REGION Network 203: DB64 DBX44.7 = PVVA Tank 8 Open Alarm
   // BWTS_ALARM_WORD_23_BIT_7
   RUNG wire#powerrail
      Contact( "1092_HMI_OP_FLAGS".CV427_428_PVVA_Alarms[8].Open )
      Coil( %DB60.DBX44.7 )
   END_RUNG
   // the same network as SCL:
   %DB60.DBX44.7 := "1092_HMI_OP_FLAGS".CV427_428_PVVA_Alarms[8].Open;
END_REGION

REGION Network 204: DB64 DBX45.0 = PVVA Tank 9 Open Alarm
   // BWTS_ALARM_WORD_23_BIT_8
   RUNG wire#powerrail
      Contact( "1092_HMI_OP_FLAGS".CV427_428_PVVA_Alarms[9].Open )
      Coil( %DB60.DBX45.0 )
   END_RUNG
   // the same network as SCL:
   %DB60.DBX45.0 := "1092_HMI_OP_FLAGS".CV427_428_PVVA_Alarms[9].Open;
END_REGION

REGION Network 205: DB64 DBX45.1 = PVVA Tank 10 Open Alarm
   // BWTS_ALARM_WORD_23_BIT_9
   RUNG wire#powerrail
      Contact( "1092_HMI_OP_FLAGS".CV427_428_PVVA_Alarms[10].Open )
      Coil( %DB60.DBX45.1 )
   END_RUNG
   // the same network as SCL:
   %DB60.DBX45.1 := "1092_HMI_OP_FLAGS".CV427_428_PVVA_Alarms[10].Open;
END_REGION

REGION Network 206: DB64 DBX45.2 = PVVA Tank 11 Open Alarm
   // BWTS_ALARM_WORD_23_BIT_10
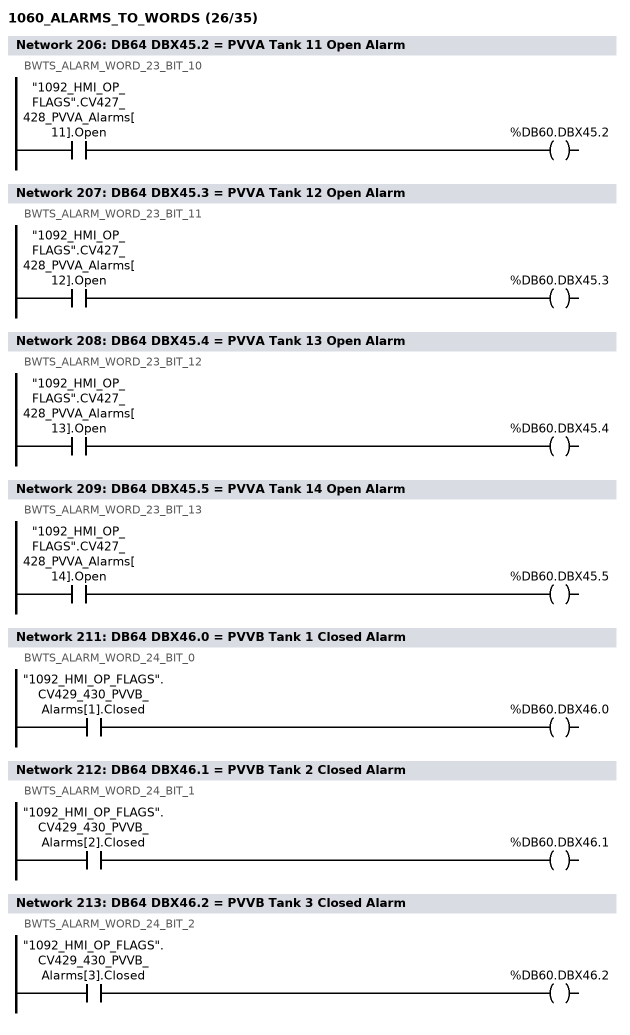
   RUNG wire#powerrail
      Contact( "1092_HMI_OP_FLAGS".CV427_428_PVVA_Alarms[11].Open )
      Coil( %DB60.DBX45.2 )
   END_RUNG
   // the same network as SCL:
   %DB60.DBX45.2 := "1092_HMI_OP_FLAGS".CV427_428_PVVA_Alarms[11].Open;
END_REGION

REGION Network 207: DB64 DBX45.3 = PVVA Tank 12 Open Alarm
   // BWTS_ALARM_WORD_23_BIT_11
   RUNG wire#powerrail
      Contact( "1092_HMI_OP_FLAGS".CV427_428_PVVA_Alarms[12].Open )
      Coil( %DB60.DBX45.3 )
   END_RUNG
   // the same network as SCL:
   %DB60.DBX45.3 := "1092_HMI_OP_FLAGS".CV427_428_PVVA_Alarms[12].Open;
END_REGION

REGION Network 208: DB64 DBX45.4 = PVVA Tank 13 Open Alarm
   // BWTS_ALARM_WORD_23_BIT_12
   RUNG wire#powerrail
      Contact( "1092_HMI_OP_FLAGS".CV427_428_PVVA_Alarms[13].Open )
      Coil( %DB60.DBX45.4 )
   END_RUNG
   // the same network as SCL:
   %DB60.DBX45.4 := "1092_HMI_OP_FLAGS".CV427_428_PVVA_Alarms[13].Open;
END_REGION

REGION Network 209: DB64 DBX45.5 = PVVA Tank 14 Open Alarm
   // BWTS_ALARM_WORD_23_BIT_13
   RUNG wire#powerrail
      Contact( "1092_HMI_OP_FLAGS".CV427_428_PVVA_Alarms[14].Open )
      Coil( %DB60.DBX45.5 )
   END_RUNG
   // the same network as SCL:
   %DB60.DBX45.5 := "1092_HMI_OP_FLAGS".CV427_428_PVVA_Alarms[14].Open;
END_REGION

REGION Network 211: DB64 DBX46.0 = PVVB Tank 1 Closed Alarm
   // BWTS_ALARM_WORD_24_BIT_0
   RUNG wire#powerrail
      Contact( "1092_HMI_OP_FLAGS".CV429_430_PVVB_Alarms[1].Closed )
      Coil( %DB60.DBX46.0 )
   END_RUNG
   // the same network as SCL:
   %DB60.DBX46.0 := "1092_HMI_OP_FLAGS".CV429_430_PVVB_Alarms[1].Closed;
END_REGION

REGION Network 212: DB64 DBX46.1 = PVVB Tank 2 Closed Alarm
   // BWTS_ALARM_WORD_24_BIT_1
   RUNG wire#powerrail
      Contact( "1092_HMI_OP_FLAGS".CV429_430_PVVB_Alarms[2].Closed )
      Coil( %DB60.DBX46.1 )
   END_RUNG
   // the same network as SCL:
   %DB60.DBX46.1 := "1092_HMI_OP_FLAGS".CV429_430_PVVB_Alarms[2].Closed;
END_REGION

REGION Network 213: DB64 DBX46.2 = PVVB Tank 3 Closed Alarm
   // BWTS_ALARM_WORD_24_BIT_2
   RUNG wire#powerrail
      Contact( "1092_HMI_OP_FLAGS".CV429_430_PVVB_Alarms[3].Closed )
      Coil( %DB60.DBX46.2 )
   END_RUNG
   // the same network as SCL:
   %DB60.DBX46.2 := "1092_HMI_OP_FLAGS".CV429_430_PVVB_Alarms[3].Closed;
END_REGION

REGION Network 214: DB64 DBX46.3 = PVVB Tank 4 Closed Alarm
   // BWTS_ALARM_WORD_24_BIT_3
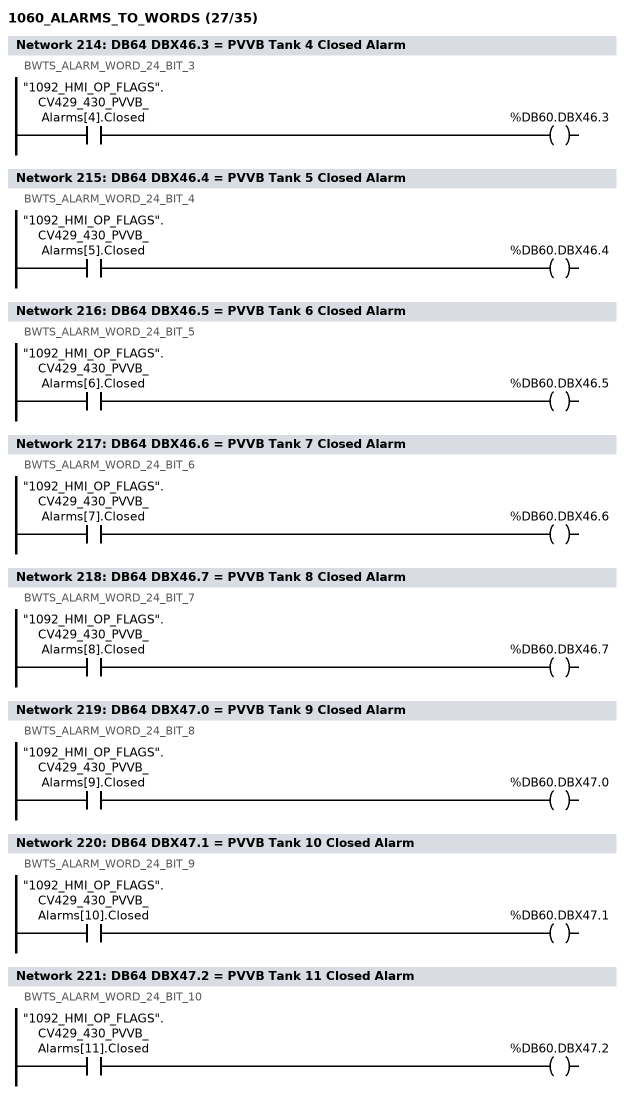
   RUNG wire#powerrail
      Contact( "1092_HMI_OP_FLAGS".CV429_430_PVVB_Alarms[4].Closed )
      Coil( %DB60.DBX46.3 )
   END_RUNG
   // the same network as SCL:
   %DB60.DBX46.3 := "1092_HMI_OP_FLAGS".CV429_430_PVVB_Alarms[4].Closed;
END_REGION

REGION Network 215: DB64 DBX46.4 = PVVB Tank 5 Closed Alarm
   // BWTS_ALARM_WORD_24_BIT_4
   RUNG wire#powerrail
      Contact( "1092_HMI_OP_FLAGS".CV429_430_PVVB_Alarms[5].Closed )
      Coil( %DB60.DBX46.4 )
   END_RUNG
   // the same network as SCL:
   %DB60.DBX46.4 := "1092_HMI_OP_FLAGS".CV429_430_PVVB_Alarms[5].Closed;
END_REGION

REGION Network 216: DB64 DBX46.5 = PVVB Tank 6 Closed Alarm
   // BWTS_ALARM_WORD_24_BIT_5
   RUNG wire#powerrail
      Contact( "1092_HMI_OP_FLAGS".CV429_430_PVVB_Alarms[6].Closed )
      Coil( %DB60.DBX46.5 )
   END_RUNG
   // the same network as SCL:
   %DB60.DBX46.5 := "1092_HMI_OP_FLAGS".CV429_430_PVVB_Alarms[6].Closed;
END_REGION

REGION Network 217: DB64 DBX46.6 = PVVB Tank 7 Closed Alarm
   // BWTS_ALARM_WORD_24_BIT_6
   RUNG wire#powerrail
      Contact( "1092_HMI_OP_FLAGS".CV429_430_PVVB_Alarms[7].Closed )
      Coil( %DB60.DBX46.6 )
   END_RUNG
   // the same network as SCL:
   %DB60.DBX46.6 := "1092_HMI_OP_FLAGS".CV429_430_PVVB_Alarms[7].Closed;
END_REGION

REGION Network 218: DB64 DBX46.7 = PVVB Tank 8 Closed Alarm
   // BWTS_ALARM_WORD_24_BIT_7
   RUNG wire#powerrail
      Contact( "1092_HMI_OP_FLAGS".CV429_430_PVVB_Alarms[8].Closed )
      Coil( %DB60.DBX46.7 )
   END_RUNG
   // the same network as SCL:
   %DB60.DBX46.7 := "1092_HMI_OP_FLAGS".CV429_430_PVVB_Alarms[8].Closed;
END_REGION

REGION Network 219: DB64 DBX47.0 = PVVB Tank 9 Closed Alarm
   // BWTS_ALARM_WORD_24_BIT_8
   RUNG wire#powerrail
      Contact( "1092_HMI_OP_FLAGS".CV429_430_PVVB_Alarms[9].Closed )
      Coil( %DB60.DBX47.0 )
   END_RUNG
   // the same network as SCL:
   %DB60.DBX47.0 := "1092_HMI_OP_FLAGS".CV429_430_PVVB_Alarms[9].Closed;
END_REGION

REGION Network 220: DB64 DBX47.1 = PVVB Tank 10 Closed Alarm
   // BWTS_ALARM_WORD_24_BIT_9
   RUNG wire#powerrail
      Contact( "1092_HMI_OP_FLAGS".CV429_430_PVVB_Alarms[10].Closed )
      Coil( %DB60.DBX47.1 )
   END_RUNG
   // the same network as SCL:
   %DB60.DBX47.1 := "1092_HMI_OP_FLAGS".CV429_430_PVVB_Alarms[10].Closed;
END_REGION

REGION Network 221: DB64 DBX47.2 = PVVB Tank 11 Closed Alarm
   // BWTS_ALARM_WORD_24_BIT_10
   RUNG wire#powerrail
      Contact( "1092_HMI_OP_FLAGS".CV429_430_PVVB_Alarms[11].Closed )
      Coil( %DB60.DBX47.2 )
   END_RUNG
   // the same network as SCL:
   %DB60.DBX47.2 := "1092_HMI_OP_FLAGS".CV429_430_PVVB_Alarms[11].Closed;
END_REGION

REGION Network 222: DB64 DBX47.3 = PVVB Tank 12 Closed Alarm
   // BWTS_ALARM_WORD_24_BIT_11
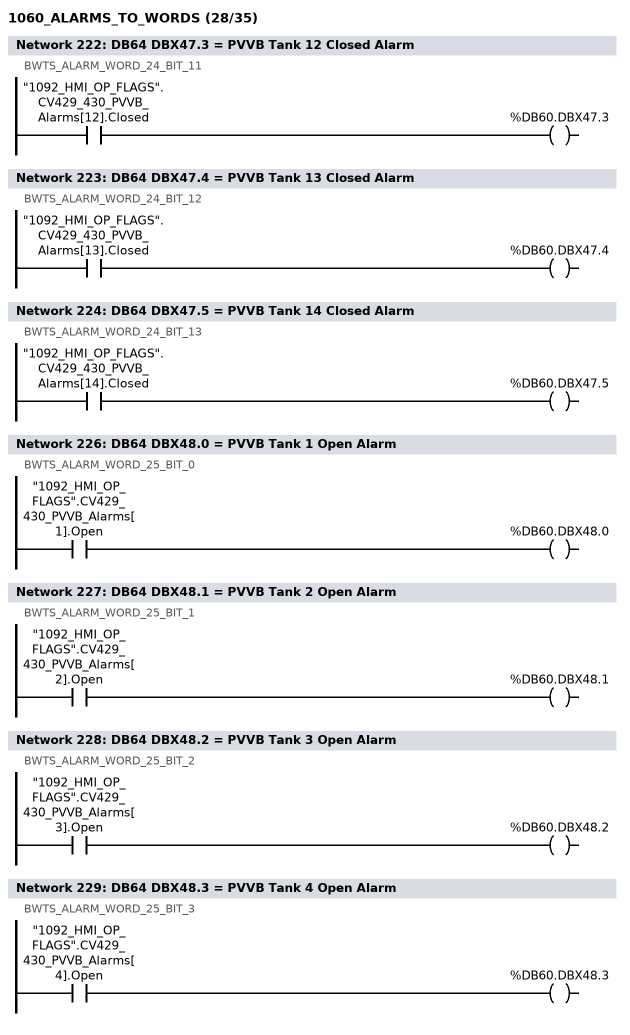
   RUNG wire#powerrail
      Contact( "1092_HMI_OP_FLAGS".CV429_430_PVVB_Alarms[12].Closed )
      Coil( %DB60.DBX47.3 )
   END_RUNG
   // the same network as SCL:
   %DB60.DBX47.3 := "1092_HMI_OP_FLAGS".CV429_430_PVVB_Alarms[12].Closed;
END_REGION

REGION Network 223: DB64 DBX47.4 = PVVB Tank 13 Closed Alarm
   // BWTS_ALARM_WORD_24_BIT_12
   RUNG wire#powerrail
      Contact( "1092_HMI_OP_FLAGS".CV429_430_PVVB_Alarms[13].Closed )
      Coil( %DB60.DBX47.4 )
   END_RUNG
   // the same network as SCL:
   %DB60.DBX47.4 := "1092_HMI_OP_FLAGS".CV429_430_PVVB_Alarms[13].Closed;
END_REGION

REGION Network 224: DB64 DBX47.5 = PVVB Tank 14 Closed Alarm
   // BWTS_ALARM_WORD_24_BIT_13
   RUNG wire#powerrail
      Contact( "1092_HMI_OP_FLAGS".CV429_430_PVVB_Alarms[14].Closed )
      Coil( %DB60.DBX47.5 )
   END_RUNG
   // the same network as SCL:
   %DB60.DBX47.5 := "1092_HMI_OP_FLAGS".CV429_430_PVVB_Alarms[14].Closed;
END_REGION

REGION Network 226: DB64 DBX48.0 = PVVB Tank 1 Open Alarm
   // BWTS_ALARM_WORD_25_BIT_0
   RUNG wire#powerrail
      Contact( "1092_HMI_OP_FLAGS".CV429_430_PVVB_Alarms[1].Open )
      Coil( %DB60.DBX48.0 )
   END_RUNG
   // the same network as SCL:
   %DB60.DBX48.0 := "1092_HMI_OP_FLAGS".CV429_430_PVVB_Alarms[1].Open;
END_REGION

REGION Network 227: DB64 DBX48.1 = PVVB Tank 2 Open Alarm
   // BWTS_ALARM_WORD_25_BIT_1
   RUNG wire#powerrail
      Contact( "1092_HMI_OP_FLAGS".CV429_430_PVVB_Alarms[2].Open )
      Coil( %DB60.DBX48.1 )
   END_RUNG
   // the same network as SCL:
   %DB60.DBX48.1 := "1092_HMI_OP_FLAGS".CV429_430_PVVB_Alarms[2].Open;
END_REGION

REGION Network 228: DB64 DBX48.2 = PVVB Tank 3 Open Alarm
   // BWTS_ALARM_WORD_25_BIT_2
   RUNG wire#powerrail
      Contact( "1092_HMI_OP_FLAGS".CV429_430_PVVB_Alarms[3].Open )
      Coil( %DB60.DBX48.2 )
   END_RUNG
   // the same network as SCL:
   %DB60.DBX48.2 := "1092_HMI_OP_FLAGS".CV429_430_PVVB_Alarms[3].Open;
END_REGION

REGION Network 229: DB64 DBX48.3 = PVVB Tank 4 Open Alarm
   // BWTS_ALARM_WORD_25_BIT_3
   RUNG wire#powerrail
      Contact( "1092_HMI_OP_FLAGS".CV429_430_PVVB_Alarms[4].Open )
      Coil( %DB60.DBX48.3 )
   END_RUNG
   // the same network as SCL:
   %DB60.DBX48.3 := "1092_HMI_OP_FLAGS".CV429_430_PVVB_Alarms[4].Open;
END_REGION

REGION Network 230: DB64 DBX48.4 = PVVB Tank 5 Open Alarm
   // BWTS_ALARM_WORD_25_BIT_4
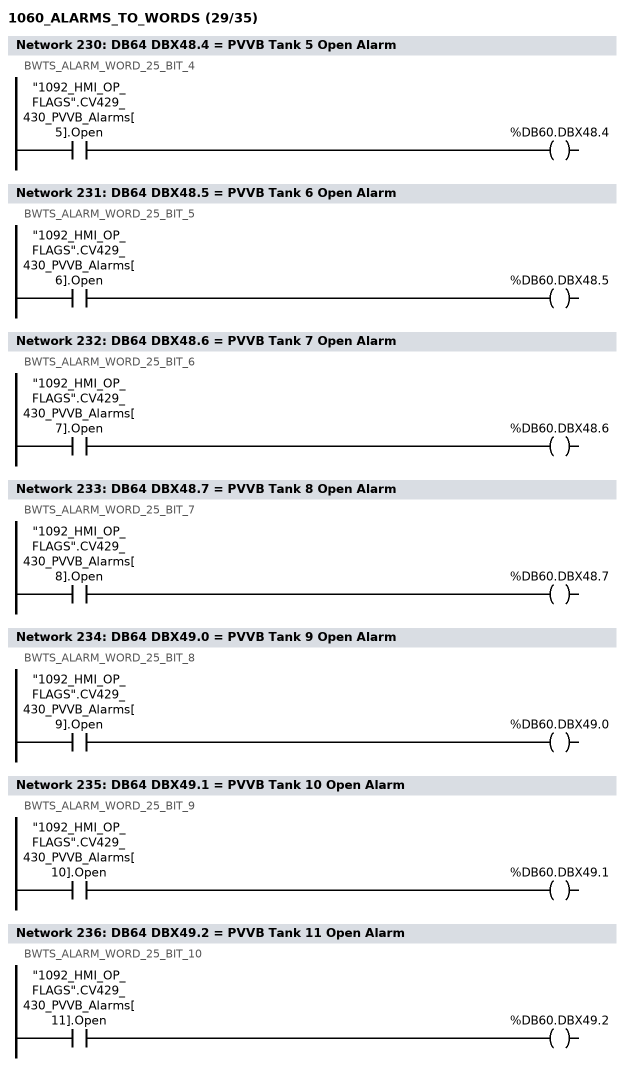
   RUNG wire#powerrail
      Contact( "1092_HMI_OP_FLAGS".CV429_430_PVVB_Alarms[5].Open )
      Coil( %DB60.DBX48.4 )
   END_RUNG
   // the same network as SCL:
   %DB60.DBX48.4 := "1092_HMI_OP_FLAGS".CV429_430_PVVB_Alarms[5].Open;
END_REGION

REGION Network 231: DB64 DBX48.5 = PVVB Tank 6 Open Alarm
   // BWTS_ALARM_WORD_25_BIT_5
   RUNG wire#powerrail
      Contact( "1092_HMI_OP_FLAGS".CV429_430_PVVB_Alarms[6].Open )
      Coil( %DB60.DBX48.5 )
   END_RUNG
   // the same network as SCL:
   %DB60.DBX48.5 := "1092_HMI_OP_FLAGS".CV429_430_PVVB_Alarms[6].Open;
END_REGION

REGION Network 232: DB64 DBX48.6 = PVVB Tank 7 Open Alarm
   // BWTS_ALARM_WORD_25_BIT_6
   RUNG wire#powerrail
      Contact( "1092_HMI_OP_FLAGS".CV429_430_PVVB_Alarms[7].Open )
      Coil( %DB60.DBX48.6 )
   END_RUNG
   // the same network as SCL:
   %DB60.DBX48.6 := "1092_HMI_OP_FLAGS".CV429_430_PVVB_Alarms[7].Open;
END_REGION

REGION Network 233: DB64 DBX48.7 = PVVB Tank 8 Open Alarm
   // BWTS_ALARM_WORD_25_BIT_7
   RUNG wire#powerrail
      Contact( "1092_HMI_OP_FLAGS".CV429_430_PVVB_Alarms[8].Open )
      Coil( %DB60.DBX48.7 )
   END_RUNG
   // the same network as SCL:
   %DB60.DBX48.7 := "1092_HMI_OP_FLAGS".CV429_430_PVVB_Alarms[8].Open;
END_REGION

REGION Network 234: DB64 DBX49.0 = PVVB Tank 9 Open Alarm
   // BWTS_ALARM_WORD_25_BIT_8
   RUNG wire#powerrail
      Contact( "1092_HMI_OP_FLAGS".CV429_430_PVVB_Alarms[9].Open )
      Coil( %DB60.DBX49.0 )
   END_RUNG
   // the same network as SCL:
   %DB60.DBX49.0 := "1092_HMI_OP_FLAGS".CV429_430_PVVB_Alarms[9].Open;
END_REGION

REGION Network 235: DB64 DBX49.1 = PVVB Tank 10 Open Alarm
   // BWTS_ALARM_WORD_25_BIT_9
   RUNG wire#powerrail
      Contact( "1092_HMI_OP_FLAGS".CV429_430_PVVB_Alarms[10].Open )
      Coil( %DB60.DBX49.1 )
   END_RUNG
   // the same network as SCL:
   %DB60.DBX49.1 := "1092_HMI_OP_FLAGS".CV429_430_PVVB_Alarms[10].Open;
END_REGION

REGION Network 236: DB64 DBX49.2 = PVVB Tank 11 Open Alarm
   // BWTS_ALARM_WORD_25_BIT_10
   RUNG wire#powerrail
      Contact( "1092_HMI_OP_FLAGS".CV429_430_PVVB_Alarms[11].Open )
      Coil( %DB60.DBX49.2 )
   END_RUNG
   // the same network as SCL:
   %DB60.DBX49.2 := "1092_HMI_OP_FLAGS".CV429_430_PVVB_Alarms[11].Open;
END_REGION

REGION Network 237: DB64 DBX49.3 = PVVB Tank 12 Open Alarm
   // BWTS_ALARM_WORD_25_BIT_11
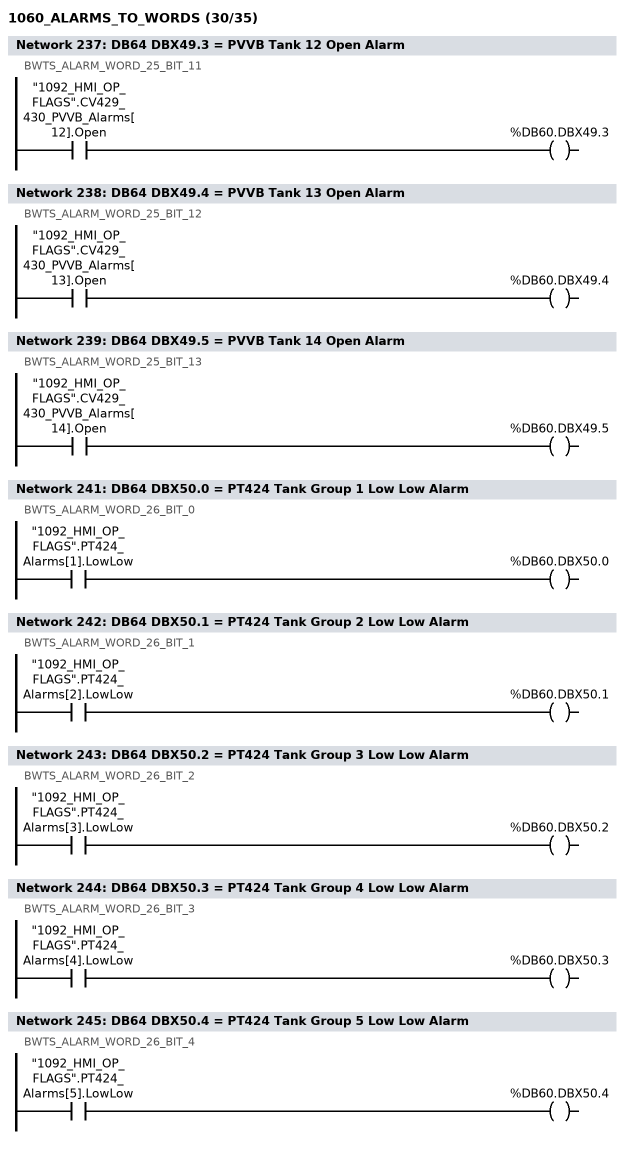
   RUNG wire#powerrail
      Contact( "1092_HMI_OP_FLAGS".CV429_430_PVVB_Alarms[12].Open )
      Coil( %DB60.DBX49.3 )
   END_RUNG
   // the same network as SCL:
   %DB60.DBX49.3 := "1092_HMI_OP_FLAGS".CV429_430_PVVB_Alarms[12].Open;
END_REGION

REGION Network 238: DB64 DBX49.4 = PVVB Tank 13 Open Alarm
   // BWTS_ALARM_WORD_25_BIT_12
   RUNG wire#powerrail
      Contact( "1092_HMI_OP_FLAGS".CV429_430_PVVB_Alarms[13].Open )
      Coil( %DB60.DBX49.4 )
   END_RUNG
   // the same network as SCL:
   %DB60.DBX49.4 := "1092_HMI_OP_FLAGS".CV429_430_PVVB_Alarms[13].Open;
END_REGION

REGION Network 239: DB64 DBX49.5 = PVVB Tank 14 Open Alarm
   // BWTS_ALARM_WORD_25_BIT_13
   RUNG wire#powerrail
      Contact( "1092_HMI_OP_FLAGS".CV429_430_PVVB_Alarms[14].Open )
      Coil( %DB60.DBX49.5 )
   END_RUNG
   // the same network as SCL:
   %DB60.DBX49.5 := "1092_HMI_OP_FLAGS".CV429_430_PVVB_Alarms[14].Open;
END_REGION

REGION Network 241: DB64 DBX50.0 = PT424 Tank Group 1 Low Low Alarm
   // BWTS_ALARM_WORD_26_BIT_0
   RUNG wire#powerrail
      Contact( "1092_HMI_OP_FLAGS".PT424_Alarms[1].LowLow )
      Coil( %DB60.DBX50.0 )
   END_RUNG
   // the same network as SCL:
   %DB60.DBX50.0 := "1092_HMI_OP_FLAGS".PT424_Alarms[1].LowLow;
END_REGION

REGION Network 242: DB64 DBX50.1 = PT424 Tank Group 2 Low Low Alarm
   // BWTS_ALARM_WORD_26_BIT_1
   RUNG wire#powerrail
      Contact( "1092_HMI_OP_FLAGS".PT424_Alarms[2].LowLow )
      Coil( %DB60.DBX50.1 )
   END_RUNG
   // the same network as SCL:
   %DB60.DBX50.1 := "1092_HMI_OP_FLAGS".PT424_Alarms[2].LowLow;
END_REGION

REGION Network 243: DB64 DBX50.2 = PT424 Tank Group 3 Low Low Alarm
   // BWTS_ALARM_WORD_26_BIT_2
   RUNG wire#powerrail
      Contact( "1092_HMI_OP_FLAGS".PT424_Alarms[3].LowLow )
      Coil( %DB60.DBX50.2 )
   END_RUNG
   // the same network as SCL:
   %DB60.DBX50.2 := "1092_HMI_OP_FLAGS".PT424_Alarms[3].LowLow;
END_REGION

REGION Network 244: DB64 DBX50.3 = PT424 Tank Group 4 Low Low Alarm
   // BWTS_ALARM_WORD_26_BIT_3
   RUNG wire#powerrail
      Contact( "1092_HMI_OP_FLAGS".PT424_Alarms[4].LowLow )
      Coil( %DB60.DBX50.3 )
   END_RUNG
   // the same network as SCL:
   %DB60.DBX50.3 := "1092_HMI_OP_FLAGS".PT424_Alarms[4].LowLow;
END_REGION

REGION Network 245: DB64 DBX50.4 = PT424 Tank Group 5 Low Low Alarm
   // BWTS_ALARM_WORD_26_BIT_4
   RUNG wire#powerrail
      Contact( "1092_HMI_OP_FLAGS".PT424_Alarms[5].LowLow )
      Coil( %DB60.DBX50.4 )
   END_RUNG
   // the same network as SCL:
   %DB60.DBX50.4 := "1092_HMI_OP_FLAGS".PT424_Alarms[5].LowLow;
END_REGION

REGION Network 246: DB64 DBX50.5 = PT424 Tank Group 6 Low Low Alarm
   // BWTS_ALARM_WORD_26_BIT_5
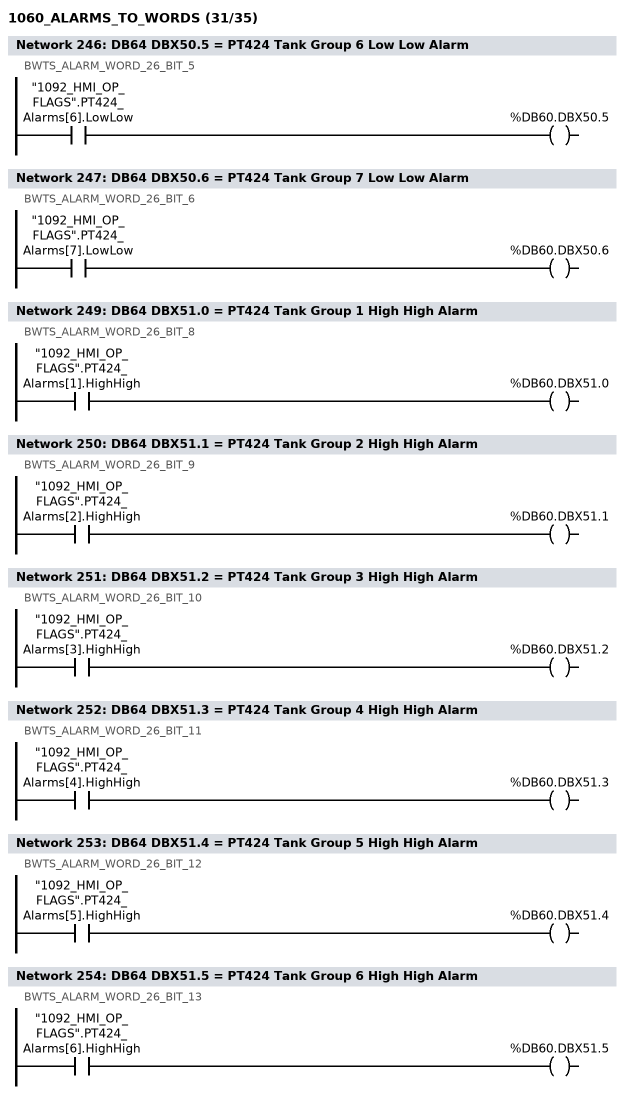
   RUNG wire#powerrail
      Contact( "1092_HMI_OP_FLAGS".PT424_Alarms[6].LowLow )
      Coil( %DB60.DBX50.5 )
   END_RUNG
   // the same network as SCL:
   %DB60.DBX50.5 := "1092_HMI_OP_FLAGS".PT424_Alarms[6].LowLow;
END_REGION

REGION Network 247: DB64 DBX50.6 = PT424 Tank Group 7 Low Low Alarm
   // BWTS_ALARM_WORD_26_BIT_6
   RUNG wire#powerrail
      Contact( "1092_HMI_OP_FLAGS".PT424_Alarms[7].LowLow )
      Coil( %DB60.DBX50.6 )
   END_RUNG
   // the same network as SCL:
   %DB60.DBX50.6 := "1092_HMI_OP_FLAGS".PT424_Alarms[7].LowLow;
END_REGION

REGION Network 249: DB64 DBX51.0 = PT424 Tank Group 1 High High Alarm
   // BWTS_ALARM_WORD_26_BIT_8
   RUNG wire#powerrail
      Contact( "1092_HMI_OP_FLAGS".PT424_Alarms[1].HighHigh )
      Coil( %DB60.DBX51.0 )
   END_RUNG
   // the same network as SCL:
   %DB60.DBX51.0 := "1092_HMI_OP_FLAGS".PT424_Alarms[1].HighHigh;
END_REGION

REGION Network 250: DB64 DBX51.1 = PT424 Tank Group 2 High High Alarm
   // BWTS_ALARM_WORD_26_BIT_9
   RUNG wire#powerrail
      Contact( "1092_HMI_OP_FLAGS".PT424_Alarms[2].HighHigh )
      Coil( %DB60.DBX51.1 )
   END_RUNG
   // the same network as SCL:
   %DB60.DBX51.1 := "1092_HMI_OP_FLAGS".PT424_Alarms[2].HighHigh;
END_REGION

REGION Network 251: DB64 DBX51.2 = PT424 Tank Group 3 High High Alarm
   // BWTS_ALARM_WORD_26_BIT_10
   RUNG wire#powerrail
      Contact( "1092_HMI_OP_FLAGS".PT424_Alarms[3].HighHigh )
      Coil( %DB60.DBX51.2 )
   END_RUNG
   // the same network as SCL:
   %DB60.DBX51.2 := "1092_HMI_OP_FLAGS".PT424_Alarms[3].HighHigh;
END_REGION

REGION Network 252: DB64 DBX51.3 = PT424 Tank Group 4 High High Alarm
   // BWTS_ALARM_WORD_26_BIT_11
   RUNG wire#powerrail
      Contact( "1092_HMI_OP_FLAGS".PT424_Alarms[4].HighHigh )
      Coil( %DB60.DBX51.3 )
   END_RUNG
   // the same network as SCL:
   %DB60.DBX51.3 := "1092_HMI_OP_FLAGS".PT424_Alarms[4].HighHigh;
END_REGION

REGION Network 253: DB64 DBX51.4 = PT424 Tank Group 5 High High Alarm
   // BWTS_ALARM_WORD_26_BIT_12
   RUNG wire#powerrail
      Contact( "1092_HMI_OP_FLAGS".PT424_Alarms[5].HighHigh )
      Coil( %DB60.DBX51.4 )
   END_RUNG
   // the same network as SCL:
   %DB60.DBX51.4 := "1092_HMI_OP_FLAGS".PT424_Alarms[5].HighHigh;
END_REGION

REGION Network 254: DB64 DBX51.5 = PT424 Tank Group 6 High High Alarm
   // BWTS_ALARM_WORD_26_BIT_13
   RUNG wire#powerrail
      Contact( "1092_HMI_OP_FLAGS".PT424_Alarms[6].HighHigh )
      Coil( %DB60.DBX51.5 )
   END_RUNG
   // the same network as SCL:
   %DB60.DBX51.5 := "1092_HMI_OP_FLAGS".PT424_Alarms[6].HighHigh;
END_REGION

REGION Network 255: DB64 DBX51.6 = PT424 Tank Group 7 High High Alarm
   // BWTS_ALARM_WORD_26_BIT_14
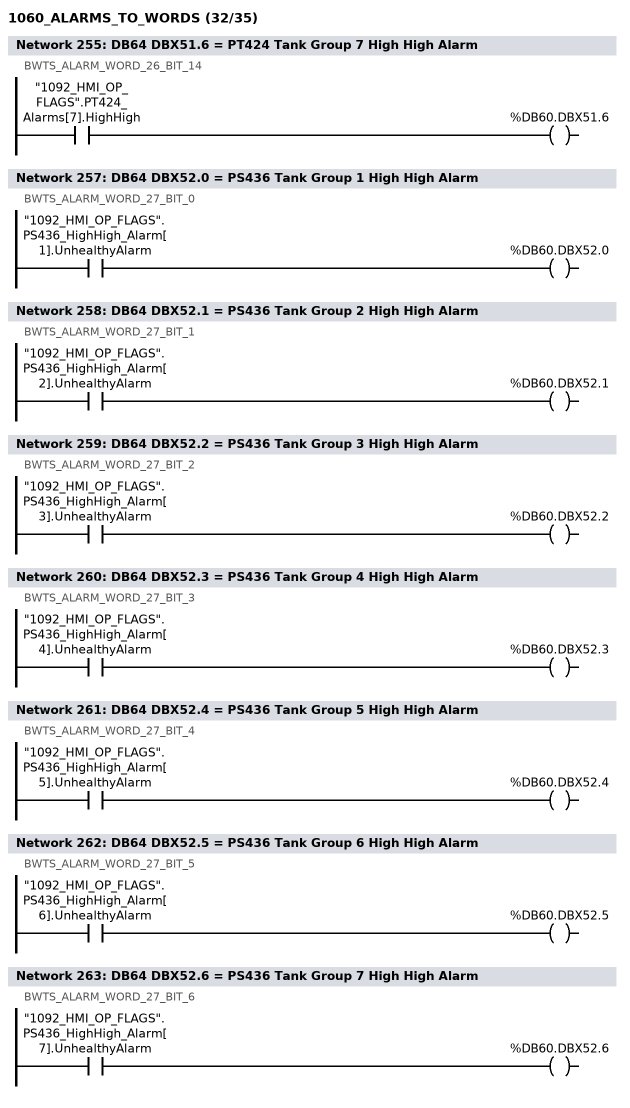
   RUNG wire#powerrail
      Contact( "1092_HMI_OP_FLAGS".PT424_Alarms[7].HighHigh )
      Coil( %DB60.DBX51.6 )
   END_RUNG
   // the same network as SCL:
   %DB60.DBX51.6 := "1092_HMI_OP_FLAGS".PT424_Alarms[7].HighHigh;
END_REGION

REGION Network 257: DB64 DBX52.0 = PS436 Tank Group 1 High High Alarm
   // BWTS_ALARM_WORD_27_BIT_0
   RUNG wire#powerrail
      Contact( "1092_HMI_OP_FLAGS".PS436_HighHigh_Alarm[1].UnhealthyAlarm )
      Coil( %DB60.DBX52.0 )
   END_RUNG
   // the same network as SCL:
   %DB60.DBX52.0 := "1092_HMI_OP_FLAGS".PS436_HighHigh_Alarm[1].UnhealthyAlarm;
END_REGION

REGION Network 258: DB64 DBX52.1 = PS436 Tank Group 2 High High Alarm
   // BWTS_ALARM_WORD_27_BIT_1
   RUNG wire#powerrail
      Contact( "1092_HMI_OP_FLAGS".PS436_HighHigh_Alarm[2].UnhealthyAlarm )
      Coil( %DB60.DBX52.1 )
   END_RUNG
   // the same network as SCL:
   %DB60.DBX52.1 := "1092_HMI_OP_FLAGS".PS436_HighHigh_Alarm[2].UnhealthyAlarm;
END_REGION

REGION Network 259: DB64 DBX52.2 = PS436 Tank Group 3 High High Alarm
   // BWTS_ALARM_WORD_27_BIT_2
   RUNG wire#powerrail
      Contact( "1092_HMI_OP_FLAGS".PS436_HighHigh_Alarm[3].UnhealthyAlarm )
      Coil( %DB60.DBX52.2 )
   END_RUNG
   // the same network as SCL:
   %DB60.DBX52.2 := "1092_HMI_OP_FLAGS".PS436_HighHigh_Alarm[3].UnhealthyAlarm;
END_REGION

REGION Network 260: DB64 DBX52.3 = PS436 Tank Group 4 High High Alarm
   // BWTS_ALARM_WORD_27_BIT_3
   RUNG wire#powerrail
      Contact( "1092_HMI_OP_FLAGS".PS436_HighHigh_Alarm[4].UnhealthyAlarm )
      Coil( %DB60.DBX52.3 )
   END_RUNG
   // the same network as SCL:
   %DB60.DBX52.3 := "1092_HMI_OP_FLAGS".PS436_HighHigh_Alarm[4].UnhealthyAlarm;
END_REGION

REGION Network 261: DB64 DBX52.4 = PS436 Tank Group 5 High High Alarm
   // BWTS_ALARM_WORD_27_BIT_4
   RUNG wire#powerrail
      Contact( "1092_HMI_OP_FLAGS".PS436_HighHigh_Alarm[5].UnhealthyAlarm )
      Coil( %DB60.DBX52.4 )
   END_RUNG
   // the same network as SCL:
   %DB60.DBX52.4 := "1092_HMI_OP_FLAGS".PS436_HighHigh_Alarm[5].UnhealthyAlarm;
END_REGION

REGION Network 262: DB64 DBX52.5 = PS436 Tank Group 6 High High Alarm
   // BWTS_ALARM_WORD_27_BIT_5
   RUNG wire#powerrail
      Contact( "1092_HMI_OP_FLAGS".PS436_HighHigh_Alarm[6].UnhealthyAlarm )
      Coil( %DB60.DBX52.5 )
   END_RUNG
   // the same network as SCL:
   %DB60.DBX52.5 := "1092_HMI_OP_FLAGS".PS436_HighHigh_Alarm[6].UnhealthyAlarm;
END_REGION

REGION Network 263: DB64 DBX52.6 = PS436 Tank Group 7 High High Alarm
   // BWTS_ALARM_WORD_27_BIT_6
   RUNG wire#powerrail
      Contact( "1092_HMI_OP_FLAGS".PS436_HighHigh_Alarm[7].UnhealthyAlarm )
      Coil( %DB60.DBX52.6 )
   END_RUNG
   // the same network as SCL:
   %DB60.DBX52.6 := "1092_HMI_OP_FLAGS".PS436_HighHigh_Alarm[7].UnhealthyAlarm;
END_REGION

REGION Network 265: DB64 DBX54.0 = PIT415 Low Low Alarm
   // BWTS_ALARM_WORD_28_BIT_0
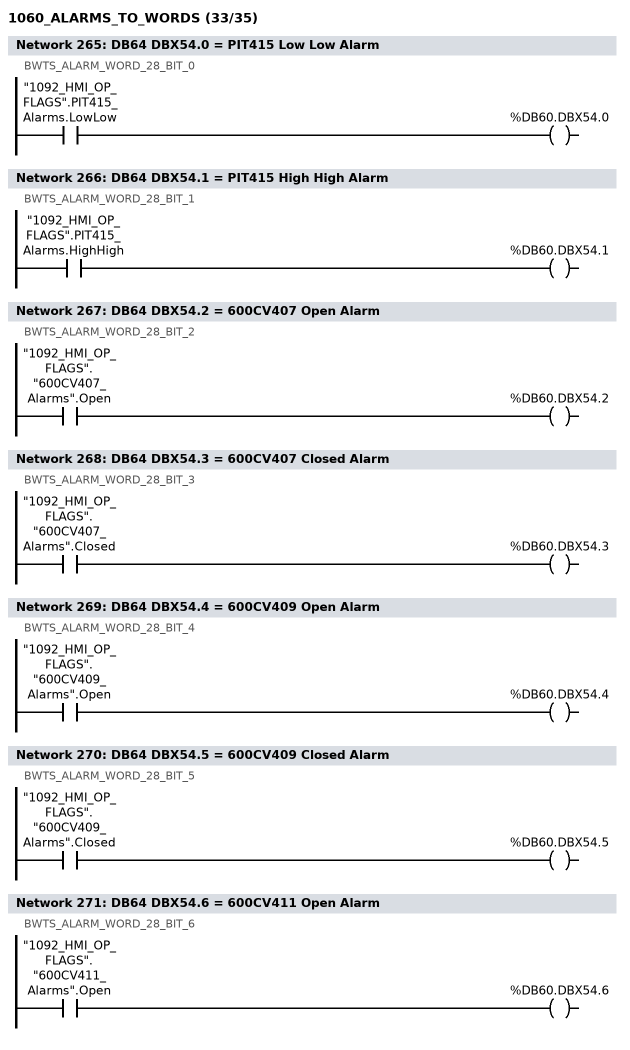
   RUNG wire#powerrail
      Contact( "1092_HMI_OP_FLAGS".PIT415_Alarms.LowLow )
      Coil( %DB60.DBX54.0 )
   END_RUNG
   // the same network as SCL:
   %DB60.DBX54.0 := "1092_HMI_OP_FLAGS".PIT415_Alarms.LowLow;
END_REGION

REGION Network 266: DB64 DBX54.1 = PIT415 High High Alarm
   // BWTS_ALARM_WORD_28_BIT_1
   RUNG wire#powerrail
      Contact( "1092_HMI_OP_FLAGS".PIT415_Alarms.HighHigh )
      Coil( %DB60.DBX54.1 )
   END_RUNG
   // the same network as SCL:
   %DB60.DBX54.1 := "1092_HMI_OP_FLAGS".PIT415_Alarms.HighHigh;
END_REGION

REGION Network 267: DB64 DBX54.2 = 600CV407 Open Alarm
   // BWTS_ALARM_WORD_28_BIT_2
   RUNG wire#powerrail
      Contact( "1092_HMI_OP_FLAGS"."600CV407_Alarms".Open )
      Coil( %DB60.DBX54.2 )
   END_RUNG
   // the same network as SCL:
   %DB60.DBX54.2 := "1092_HMI_OP_FLAGS"."600CV407_Alarms".Open;
END_REGION

REGION Network 268: DB64 DBX54.3 = 600CV407 Closed Alarm
   // BWTS_ALARM_WORD_28_BIT_3
   RUNG wire#powerrail
      Contact( "1092_HMI_OP_FLAGS"."600CV407_Alarms".Closed )
      Coil( %DB60.DBX54.3 )
   END_RUNG
   // the same network as SCL:
   %DB60.DBX54.3 := "1092_HMI_OP_FLAGS"."600CV407_Alarms".Closed;
END_REGION

REGION Network 269: DB64 DBX54.4 = 600CV409 Open Alarm
   // BWTS_ALARM_WORD_28_BIT_4
   RUNG wire#powerrail
      Contact( "1092_HMI_OP_FLAGS"."600CV409_Alarms".Open )
      Coil( %DB60.DBX54.4 )
   END_RUNG
   // the same network as SCL:
   %DB60.DBX54.4 := "1092_HMI_OP_FLAGS"."600CV409_Alarms".Open;
END_REGION

REGION Network 270: DB64 DBX54.5 = 600CV409 Closed Alarm
   // BWTS_ALARM_WORD_28_BIT_5
   RUNG wire#powerrail
      Contact( "1092_HMI_OP_FLAGS"."600CV409_Alarms".Closed )
      Coil( %DB60.DBX54.5 )
   END_RUNG
   // the same network as SCL:
   %DB60.DBX54.5 := "1092_HMI_OP_FLAGS"."600CV409_Alarms".Closed;
END_REGION

REGION Network 271: DB64 DBX54.6 = 600CV411 Open Alarm
   // BWTS_ALARM_WORD_28_BIT_6
   RUNG wire#powerrail
      Contact( "1092_HMI_OP_FLAGS"."600CV411_Alarms".Open )
      Coil( %DB60.DBX54.6 )
   END_RUNG
   // the same network as SCL:
   %DB60.DBX54.6 := "1092_HMI_OP_FLAGS"."600CV411_Alarms".Open;
END_REGION

REGION Network 272: DB64 DBX54.7 = 600CV411 Closed Alarm
   // BWTS_ALARM_WORD_28_BIT_7